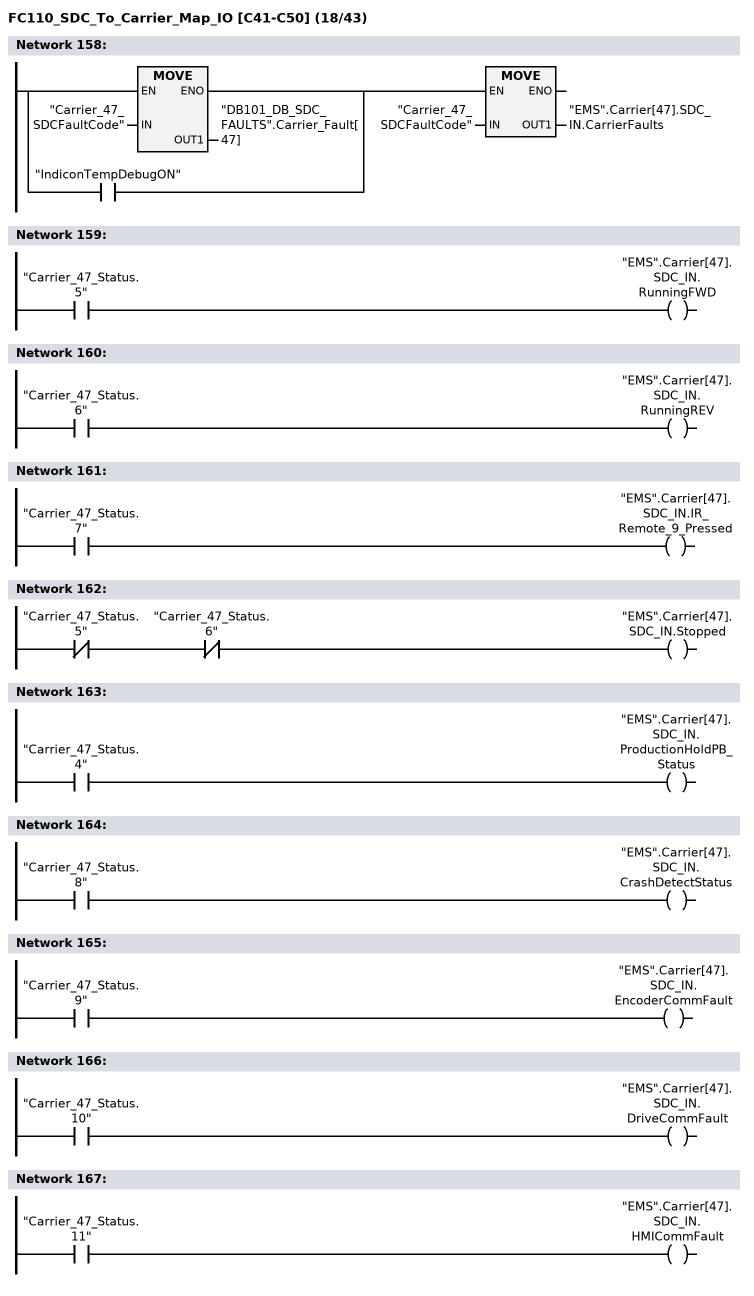
   RUNG wire#powerrail
      Move(in := "Carrier_47_SDCFaultCode", out1 => "DB101_DB_SDC_FAULTS".Carrier_Fault[47])
      wire#w1
      Move(in := "Carrier_47_SDCFaultCode", out1 => "EMS".Carrier[47].SDC_IN.CarrierFaults)
   END_RUNG
   RUNG wire#powerrail
      Contact( "IndiconTempDebugON" )
   END_RUNG wire#w1
   // the same network as SCL:
   "DB101_DB_SDC_FAULTS".Carrier_Fault[47] := "Carrier_47_SDCFaultCode";
   IF TRUE OR "IndiconTempDebugON" THEN
       "EMS".Carrier[47].SDC_IN.CarrierFaults := "Carrier_47_SDCFaultCode";
   END_IF;
END_REGION

REGION Network 159
   RUNG wire#powerrail
      Contact( "Carrier_47_Status.5" )
      Coil( "EMS".Carrier[47].SDC_IN.RunningFWD )
   END_RUNG
   // the same network as SCL:
   "EMS".Carrier[47].SDC_IN.RunningFWD := "Carrier_47_Status.5";
END_REGION

REGION Network 160
   RUNG wire#powerrail
      Contact( "Carrier_47_Status.6" )
      Coil( "EMS".Carrier[47].SDC_IN.RunningREV )
   END_RUNG
   // the same network as SCL:
   "EMS".Carrier[47].SDC_IN.RunningREV := "Carrier_47_Status.6";
END_REGION

REGION Network 161
   RUNG wire#powerrail
      Contact( "Carrier_47_Status.7" )
      Coil( "EMS".Carrier[47].SDC_IN.IR_Remote_9_Pressed )
   END_RUNG
   // the same network as SCL:
   "EMS".Carrier[47].SDC_IN.IR_Remote_9_Pressed := "Carrier_47_Status.7";
END_REGION

REGION Network 162
   RUNG wire#powerrail
      I_Contact( "Carrier_47_Status.5" )
      I_Contact( "Carrier_47_Status.6" )
      Coil( "EMS".Carrier[47].SDC_IN.Stopped )
   END_RUNG
   // the same network as SCL:
   "EMS".Carrier[47].SDC_IN.Stopped := NOT "Carrier_47_Status.5" AND NOT "Carrier_47_Status.6";
END_REGION

REGION Network 163
   RUNG wire#powerrail
      Contact( "Carrier_47_Status.4" )
      Coil( "EMS".Carrier[47].SDC_IN.ProductionHoldPB_Status )
   END_RUNG
   // the same network as SCL:
   "EMS".Carrier[47].SDC_IN.ProductionHoldPB_Status := "Carrier_47_Status.4";
END_REGION

REGION Network 164
   RUNG wire#powerrail
      Contact( "Carrier_47_Status.8" )
      Coil( "EMS".Carrier[47].SDC_IN.CrashDetectStatus )
   END_RUNG
   // the same network as SCL:
   "EMS".Carrier[47].SDC_IN.CrashDetectStatus := "Carrier_47_Status.8";
END_REGION

REGION Network 165
   RUNG wire#powerrail
      Contact( "Carrier_47_Status.9" )
      Coil( "EMS".Carrier[47].SDC_IN.EncoderCommFault )
   END_RUNG
   // the same network as SCL:
   "EMS".Carrier[47].SDC_IN.EncoderCommFault := "Carrier_47_Status.9";
END_REGION

REGION Network 166
   RUNG wire#powerrail
      Contact( "Carrier_47_Status.10" )
      Coil( "EMS".Carrier[47].SDC_IN.DriveCommFault )
   END_RUNG
   // the same network as SCL:
   "EMS".Carrier[47].SDC_IN.DriveCommFault := "Carrier_47_Status.10";
END_REGION

REGION Network 167
   RUNG wire#powerrail
      Contact( "Carrier_47_Status.11" )
      Coil( "EMS".Carrier[47].SDC_IN.HMICommFault )
   END_RUNG
   // the same network as SCL:
   "EMS".Carrier[47].SDC_IN.HMICommFault := "Carrier_47_Status.11";
END_REGION

REGION Network 168
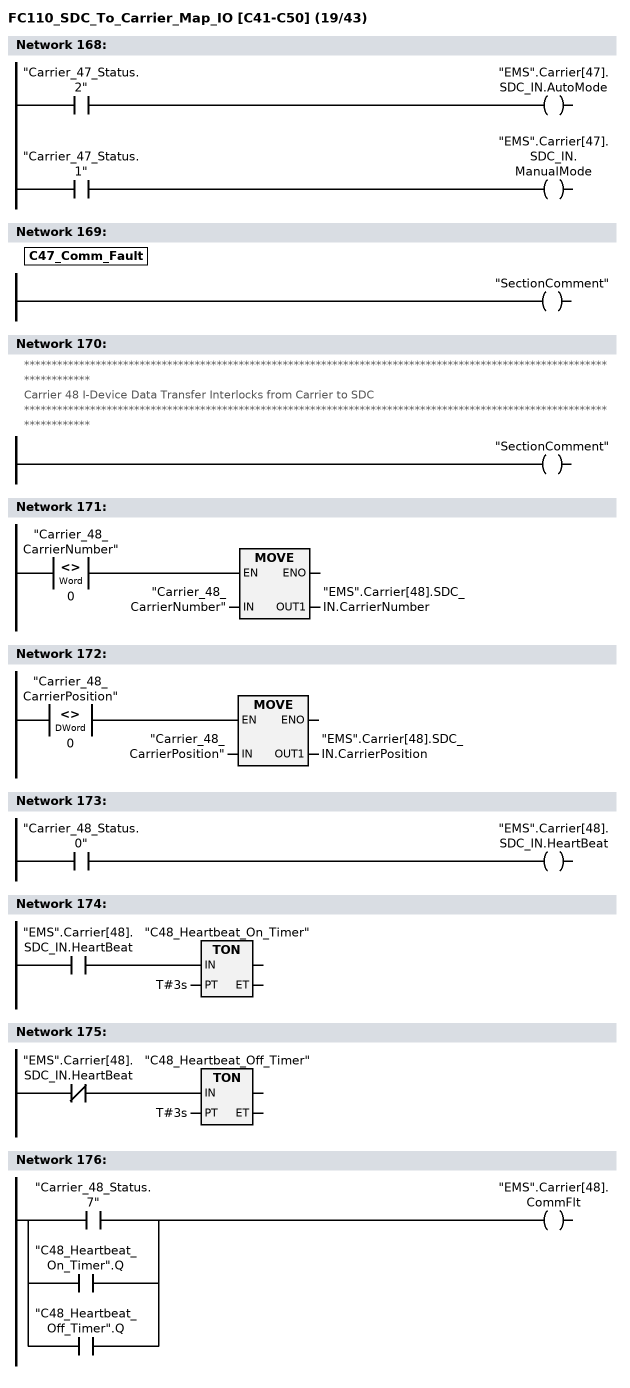
   RUNG wire#powerrail
      Contact( "Carrier_47_Status.2" )
      Coil( "EMS".Carrier[47].SDC_IN.AutoMode )
   END_RUNG
   RUNG wire#powerrail
      Contact( "Carrier_47_Status.1" )
      Coil( "EMS".Carrier[47].SDC_IN.ManualMode )
   END_RUNG
   // the same network as SCL:
   "EMS".Carrier[47].SDC_IN.AutoMode := "Carrier_47_Status.2";
   "EMS".Carrier[47].SDC_IN.ManualMode := "Carrier_47_Status.1";
END_REGION

REGION Network 169
   Label( C47_Comm_Fault )
   RUNG wire#powerrail
      Coil( "SectionComment" )
   END_RUNG
   // the same network as SCL:
   C47_Comm_Fault:
   "SectionComment" := TRUE;
END_REGION

REGION Network 170
   // **********************************************************************************************************************
   // 
   // Carrier 48 I-Device Data Transfer Interlocks from Carrier to SDC
   // 
   // **********************************************************************************************************************
   RUNG wire#powerrail
      Coil( "SectionComment" )
   END_RUNG
   // the same network as SCL:
   "SectionComment" := TRUE;
END_REGION

REGION Network 171
   RUNG wire#powerrail
      { S7_Templates := "SrcType := Word" } NE_Contact(in1 := "Carrier_48_CarrierNumber", in2 := 0)
      Move(in := "Carrier_48_CarrierNumber", out1 => "EMS".Carrier[48].SDC_IN.CarrierNumber)
   END_RUNG
   // the same network as SCL:
   IF "Carrier_48_CarrierNumber" <> 0 THEN
       "EMS".Carrier[48].SDC_IN.CarrierNumber := "Carrier_48_CarrierNumber";
   END_IF;
END_REGION

REGION Network 172
   RUNG wire#powerrail
      { S7_Templates := "SrcType := DWord" } NE_Contact(in1 := "Carrier_48_CarrierPosition", in2 := 0)
      Move(in := "Carrier_48_CarrierPosition", out1 => "EMS".Carrier[48].SDC_IN.CarrierPosition)
   END_RUNG
   // the same network as SCL:
   IF "Carrier_48_CarrierPosition" <> 0 THEN
       "EMS".Carrier[48].SDC_IN.CarrierPosition := "Carrier_48_CarrierPosition";
   END_IF;
END_REGION

REGION Network 173
   RUNG wire#powerrail
      Contact( "Carrier_48_Status.0" )
      Coil( "EMS".Carrier[48].SDC_IN.HeartBeat )
   END_RUNG
   // the same network as SCL:
   "EMS".Carrier[48].SDC_IN.HeartBeat := "Carrier_48_Status.0";
END_REGION

REGION Network 174
   "C48_Heartbeat_On_Timer".TON(IN := "EMS".Carrier[48].SDC_IN.HeartBeat, PT := T#3s);
END_REGION

REGION Network 175
   "C48_Heartbeat_Off_Timer".TON(IN := NOT "EMS".Carrier[48].SDC_IN.HeartBeat, PT := T#3s);
END_REGION

REGION Network 176
   RUNG wire#powerrail
      Contact( "Carrier_48_Status.7" )
      wire#w1
      Coil( "EMS".Carrier[48].CommFlt )
   END_RUNG
   RUNG wire#powerrail
      Contact( "C48_Heartbeat_On_Timer".Q )
   END_RUNG wire#w1
   RUNG wire#powerrail
      Contact( "C48_Heartbeat_Off_Timer".Q )
   END_RUNG wire#w1
   // the same network as SCL:
   "EMS".Carrier[48].CommFlt := "Carrier_48_Status.7" OR "C48_Heartbeat_On_Timer".Q OR "C48_Heartbeat_Off_Timer".Q;
END_REGION

REGION Network 177
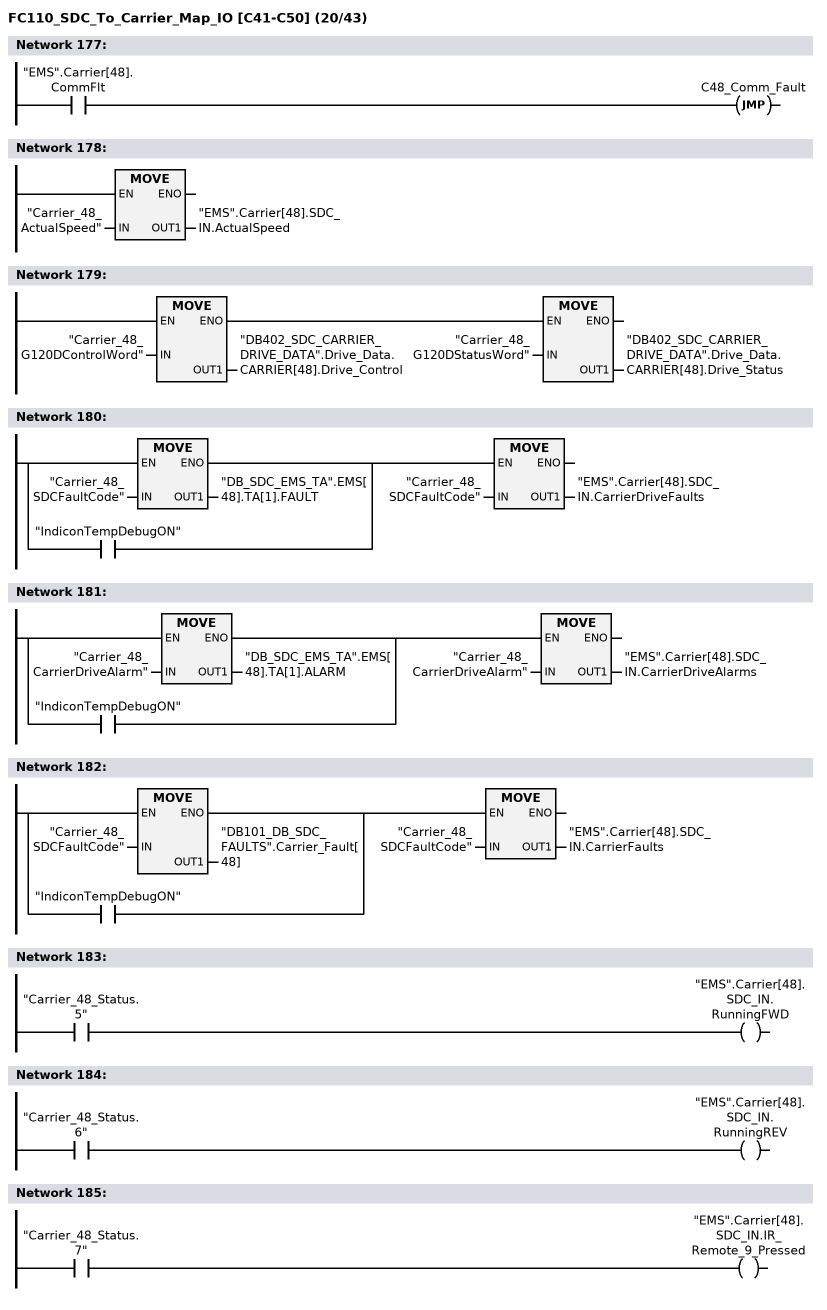
   RUNG wire#powerrail
      Contact( "EMS".Carrier[48].CommFlt )
      JumpCoil( C48_Comm_Fault )
   END_RUNG
   // the same network as SCL:
   IF "EMS".Carrier[48].CommFlt THEN GOTO C48_Comm_Fault; END_IF;
END_REGION

REGION Network 178
   RUNG wire#powerrail
      Move(in := "Carrier_48_ActualSpeed", out1 => "EMS".Carrier[48].SDC_IN.ActualSpeed)
   END_RUNG
   // the same network as SCL:
   "EMS".Carrier[48].SDC_IN.ActualSpeed := "Carrier_48_ActualSpeed";
END_REGION

REGION Network 179
   RUNG wire#powerrail
      Move(in := "Carrier_48_G120DControlWord", out1 => "DB402_SDC_CARRIER_DRIVE_DATA".Drive_Data.CARRIER[48].Drive_Control)
      Move(in := "Carrier_48_G120DStatusWord", out1 => "DB402_SDC_CARRIER_DRIVE_DATA".Drive_Data.CARRIER[48].Drive_Status)
   END_RUNG
   // the same network as SCL:
   "DB402_SDC_CARRIER_DRIVE_DATA".Drive_Data.CARRIER[48].Drive_Control := "Carrier_48_G120DControlWord";
   "DB402_SDC_CARRIER_DRIVE_DATA".Drive_Data.CARRIER[48].Drive_Status := "Carrier_48_G120DStatusWord";
END_REGION

REGION Network 180
   RUNG wire#powerrail
      Move(in := "Carrier_48_SDCFaultCode", out1 => "DB_SDC_EMS_TA".EMS[48].TA[1].FAULT)
      wire#w1
      Move(in := "Carrier_48_SDCFaultCode", out1 => "EMS".Carrier[48].SDC_IN.CarrierDriveFaults)
   END_RUNG
   RUNG wire#powerrail
      Contact( "IndiconTempDebugON" )
   END_RUNG wire#w1
   // the same network as SCL:
   "DB_SDC_EMS_TA".EMS[48].TA[1].FAULT := "Carrier_48_SDCFaultCode";
   IF TRUE OR "IndiconTempDebugON" THEN
       "EMS".Carrier[48].SDC_IN.CarrierDriveFaults := "Carrier_48_SDCFaultCode";
   END_IF;
END_REGION

REGION Network 181
   RUNG wire#powerrail
      Move(in := "Carrier_48_CarrierDriveAlarm", out1 => "DB_SDC_EMS_TA".EMS[48].TA[1].ALARM)
      wire#w1
      Move(in := "Carrier_48_CarrierDriveAlarm", out1 => "EMS".Carrier[48].SDC_IN.CarrierDriveAlarms)
   END_RUNG
   RUNG wire#powerrail
      Contact( "IndiconTempDebugON" )
   END_RUNG wire#w1
   // the same network as SCL:
   "DB_SDC_EMS_TA".EMS[48].TA[1].ALARM := "Carrier_48_CarrierDriveAlarm";
   IF TRUE OR "IndiconTempDebugON" THEN
       "EMS".Carrier[48].SDC_IN.CarrierDriveAlarms := "Carrier_48_CarrierDriveAlarm";
   END_IF;
END_REGION

REGION Network 182
   RUNG wire#powerrail
      Move(in := "Carrier_48_SDCFaultCode", out1 => "DB101_DB_SDC_FAULTS".Carrier_Fault[48])
      wire#w1
      Move(in := "Carrier_48_SDCFaultCode", out1 => "EMS".Carrier[48].SDC_IN.CarrierFaults)
   END_RUNG
   RUNG wire#powerrail
      Contact( "IndiconTempDebugON" )
   END_RUNG wire#w1
   // the same network as SCL:
   "DB101_DB_SDC_FAULTS".Carrier_Fault[48] := "Carrier_48_SDCFaultCode";
   IF TRUE OR "IndiconTempDebugON" THEN
       "EMS".Carrier[48].SDC_IN.CarrierFaults := "Carrier_48_SDCFaultCode";
   END_IF;
END_REGION

REGION Network 183
   RUNG wire#powerrail
      Contact( "Carrier_48_Status.5" )
      Coil( "EMS".Carrier[48].SDC_IN.RunningFWD )
   END_RUNG
   // the same network as SCL:
   "EMS".Carrier[48].SDC_IN.RunningFWD := "Carrier_48_Status.5";
END_REGION

REGION Network 184
   RUNG wire#powerrail
      Contact( "Carrier_48_Status.6" )
      Coil( "EMS".Carrier[48].SDC_IN.RunningREV )
   END_RUNG
   // the same network as SCL:
   "EMS".Carrier[48].SDC_IN.RunningREV := "Carrier_48_Status.6";
END_REGION

REGION Network 185
   RUNG wire#powerrail
      Contact( "Carrier_48_Status.7" )
      Coil( "EMS".Carrier[48].SDC_IN.IR_Remote_9_Pressed )
   END_RUNG
   // the same network as SCL:
   "EMS".Carrier[48].SDC_IN.IR_Remote_9_Pressed := "Carrier_48_Status.7";
END_REGION

REGION Network 186
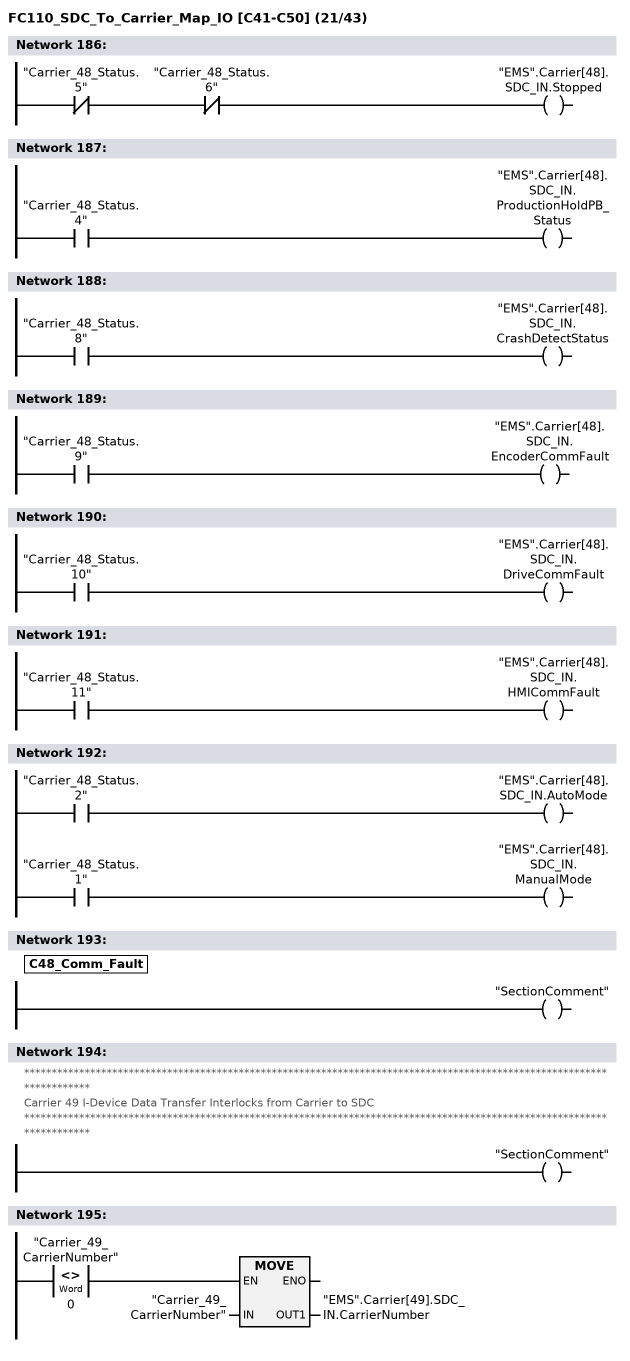
   RUNG wire#powerrail
      I_Contact( "Carrier_48_Status.5" )
      I_Contact( "Carrier_48_Status.6" )
      Coil( "EMS".Carrier[48].SDC_IN.Stopped )
   END_RUNG
   // the same network as SCL:
   "EMS".Carrier[48].SDC_IN.Stopped := NOT "Carrier_48_Status.5" AND NOT "Carrier_48_Status.6";
END_REGION

REGION Network 187
   RUNG wire#powerrail
      Contact( "Carrier_48_Status.4" )
      Coil( "EMS".Carrier[48].SDC_IN.ProductionHoldPB_Status )
   END_RUNG
   // the same network as SCL:
   "EMS".Carrier[48].SDC_IN.ProductionHoldPB_Status := "Carrier_48_Status.4";
END_REGION

REGION Network 188
   RUNG wire#powerrail
      Contact( "Carrier_48_Status.8" )
      Coil( "EMS".Carrier[48].SDC_IN.CrashDetectStatus )
   END_RUNG
   // the same network as SCL:
   "EMS".Carrier[48].SDC_IN.CrashDetectStatus := "Carrier_48_Status.8";
END_REGION

REGION Network 189
   RUNG wire#powerrail
      Contact( "Carrier_48_Status.9" )
      Coil( "EMS".Carrier[48].SDC_IN.EncoderCommFault )
   END_RUNG
   // the same network as SCL:
   "EMS".Carrier[48].SDC_IN.EncoderCommFault := "Carrier_48_Status.9";
END_REGION

REGION Network 190
   RUNG wire#powerrail
      Contact( "Carrier_48_Status.10" )
      Coil( "EMS".Carrier[48].SDC_IN.DriveCommFault )
   END_RUNG
   // the same network as SCL:
   "EMS".Carrier[48].SDC_IN.DriveCommFault := "Carrier_48_Status.10";
END_REGION

REGION Network 191
   RUNG wire#powerrail
      Contact( "Carrier_48_Status.11" )
      Coil( "EMS".Carrier[48].SDC_IN.HMICommFault )
   END_RUNG
   // the same network as SCL:
   "EMS".Carrier[48].SDC_IN.HMICommFault := "Carrier_48_Status.11";
END_REGION

REGION Network 192
   RUNG wire#powerrail
      Contact( "Carrier_48_Status.2" )
      Coil( "EMS".Carrier[48].SDC_IN.AutoMode )
   END_RUNG
   RUNG wire#powerrail
      Contact( "Carrier_48_Status.1" )
      Coil( "EMS".Carrier[48].SDC_IN.ManualMode )
   END_RUNG
   // the same network as SCL:
   "EMS".Carrier[48].SDC_IN.AutoMode := "Carrier_48_Status.2";
   "EMS".Carrier[48].SDC_IN.ManualMode := "Carrier_48_Status.1";
END_REGION

REGION Network 193
   Label( C48_Comm_Fault )
   RUNG wire#powerrail
      Coil( "SectionComment" )
   END_RUNG
   // the same network as SCL:
   C48_Comm_Fault:
   "SectionComment" := TRUE;
END_REGION

REGION Network 194
   // **********************************************************************************************************************
   // 
   // Carrier 49 I-Device Data Transfer Interlocks from Carrier to SDC
   // 
   // **********************************************************************************************************************
   RUNG wire#powerrail
      Coil( "SectionComment" )
   END_RUNG
   // the same network as SCL:
   "SectionComment" := TRUE;
END_REGION

REGION Network 195
   RUNG wire#powerrail
      { S7_Templates := "SrcType := Word" } NE_Contact(in1 := "Carrier_49_CarrierNumber", in2 := 0)
      Move(in := "Carrier_49_CarrierNumber", out1 => "EMS".Carrier[49].SDC_IN.CarrierNumber)
   END_RUNG
   // the same network as SCL:
   IF "Carrier_49_CarrierNumber" <> 0 THEN
       "EMS".Carrier[49].SDC_IN.CarrierNumber := "Carrier_49_CarrierNumber";
   END_IF;
END_REGION

REGION Network 196
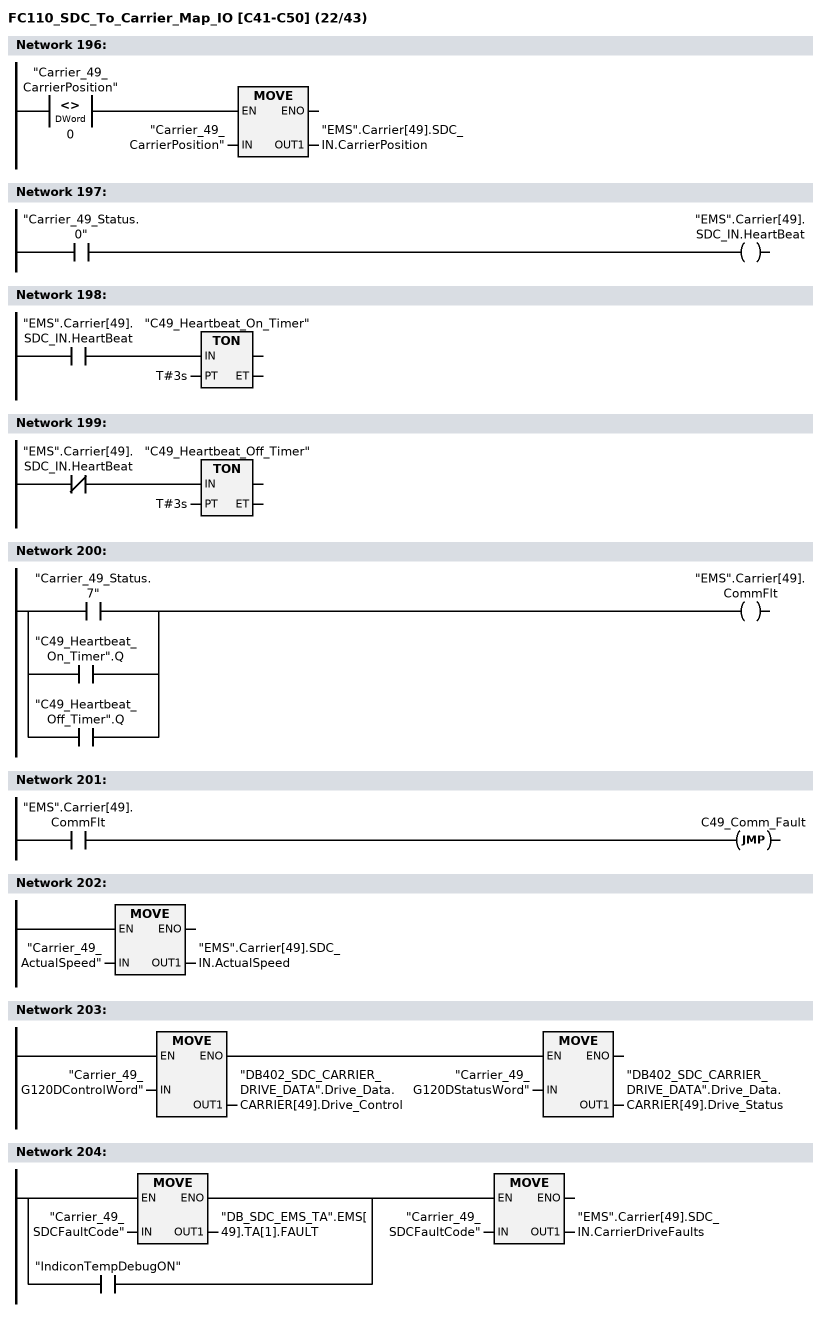
   RUNG wire#powerrail
      { S7_Templates := "SrcType := DWord" } NE_Contact(in1 := "Carrier_49_CarrierPosition", in2 := 0)
      Move(in := "Carrier_49_CarrierPosition", out1 => "EMS".Carrier[49].SDC_IN.CarrierPosition)
   END_RUNG
   // the same network as SCL:
   IF "Carrier_49_CarrierPosition" <> 0 THEN
       "EMS".Carrier[49].SDC_IN.CarrierPosition := "Carrier_49_CarrierPosition";
   END_IF;
END_REGION

REGION Network 197
   RUNG wire#powerrail
      Contact( "Carrier_49_Status.0" )
      Coil( "EMS".Carrier[49].SDC_IN.HeartBeat )
   END_RUNG
   // the same network as SCL:
   "EMS".Carrier[49].SDC_IN.HeartBeat := "Carrier_49_Status.0";
END_REGION

REGION Network 198
   "C49_Heartbeat_On_Timer".TON(IN := "EMS".Carrier[49].SDC_IN.HeartBeat, PT := T#3s);
END_REGION

REGION Network 199
   "C49_Heartbeat_Off_Timer".TON(IN := NOT "EMS".Carrier[49].SDC_IN.HeartBeat, PT := T#3s);
END_REGION

REGION Network 200
   RUNG wire#powerrail
      Contact( "Carrier_49_Status.7" )
      wire#w1
      Coil( "EMS".Carrier[49].CommFlt )
   END_RUNG
   RUNG wire#powerrail
      Contact( "C49_Heartbeat_On_Timer".Q )
   END_RUNG wire#w1
   RUNG wire#powerrail
      Contact( "C49_Heartbeat_Off_Timer".Q )
   END_RUNG wire#w1
   // the same network as SCL:
   "EMS".Carrier[49].CommFlt := "Carrier_49_Status.7" OR "C49_Heartbeat_On_Timer".Q OR "C49_Heartbeat_Off_Timer".Q;
END_REGION

REGION Network 201
   RUNG wire#powerrail
      Contact( "EMS".Carrier[49].CommFlt )
      JumpCoil( C49_Comm_Fault )
   END_RUNG
   // the same network as SCL:
   IF "EMS".Carrier[49].CommFlt THEN GOTO C49_Comm_Fault; END_IF;
END_REGION

REGION Network 202
   RUNG wire#powerrail
      Move(in := "Carrier_49_ActualSpeed", out1 => "EMS".Carrier[49].SDC_IN.ActualSpeed)
   END_RUNG
   // the same network as SCL:
   "EMS".Carrier[49].SDC_IN.ActualSpeed := "Carrier_49_ActualSpeed";
END_REGION

REGION Network 203
   RUNG wire#powerrail
      Move(in := "Carrier_49_G120DControlWord", out1 => "DB402_SDC_CARRIER_DRIVE_DATA".Drive_Data.CARRIER[49].Drive_Control)
      Move(in := "Carrier_49_G120DStatusWord", out1 => "DB402_SDC_CARRIER_DRIVE_DATA".Drive_Data.CARRIER[49].Drive_Status)
   END_RUNG
   // the same network as SCL:
   "DB402_SDC_CARRIER_DRIVE_DATA".Drive_Data.CARRIER[49].Drive_Control := "Carrier_49_G120DControlWord";
   "DB402_SDC_CARRIER_DRIVE_DATA".Drive_Data.CARRIER[49].Drive_Status := "Carrier_49_G120DStatusWord";
END_REGION

REGION Network 204
   RUNG wire#powerrail
      Move(in := "Carrier_49_SDCFaultCode", out1 => "DB_SDC_EMS_TA".EMS[49].TA[1].FAULT)
      wire#w1
      Move(in := "Carrier_49_SDCFaultCode", out1 => "EMS".Carrier[49].SDC_IN.CarrierDriveFaults)
   END_RUNG
   RUNG wire#powerrail
      Contact( "IndiconTempDebugON" )
   END_RUNG wire#w1
   // the same network as SCL:
   "DB_SDC_EMS_TA".EMS[49].TA[1].FAULT := "Carrier_49_SDCFaultCode";
   IF TRUE OR "IndiconTempDebugON" THEN
       "EMS".Carrier[49].SDC_IN.CarrierDriveFaults := "Carrier_49_SDCFaultCode";
   END_IF;
END_REGION

REGION Network 205
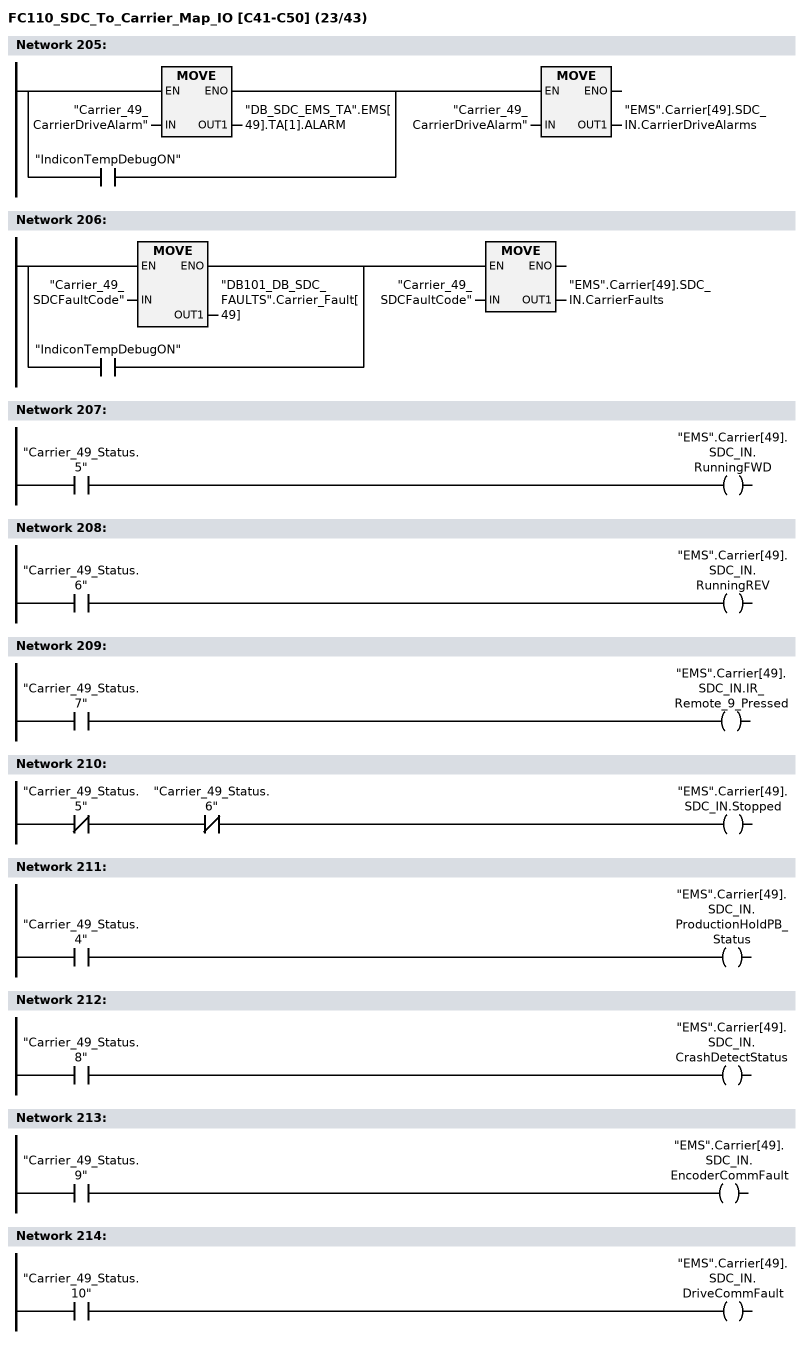
   RUNG wire#powerrail
      Move(in := "Carrier_49_CarrierDriveAlarm", out1 => "DB_SDC_EMS_TA".EMS[49].TA[1].ALARM)
      wire#w1
      Move(in := "Carrier_49_CarrierDriveAlarm", out1 => "EMS".Carrier[49].SDC_IN.CarrierDriveAlarms)
   END_RUNG
   RUNG wire#powerrail
      Contact( "IndiconTempDebugON" )
   END_RUNG wire#w1
   // the same network as SCL:
   "DB_SDC_EMS_TA".EMS[49].TA[1].ALARM := "Carrier_49_CarrierDriveAlarm";
   IF TRUE OR "IndiconTempDebugON" THEN
       "EMS".Carrier[49].SDC_IN.CarrierDriveAlarms := "Carrier_49_CarrierDriveAlarm";
   END_IF;
END_REGION

REGION Network 206
   RUNG wire#powerrail
      Move(in := "Carrier_49_SDCFaultCode", out1 => "DB101_DB_SDC_FAULTS".Carrier_Fault[49])
      wire#w1
      Move(in := "Carrier_49_SDCFaultCode", out1 => "EMS".Carrier[49].SDC_IN.CarrierFaults)
   END_RUNG
   RUNG wire#powerrail
      Contact( "IndiconTempDebugON" )
   END_RUNG wire#w1
   // the same network as SCL:
   "DB101_DB_SDC_FAULTS".Carrier_Fault[49] := "Carrier_49_SDCFaultCode";
   IF TRUE OR "IndiconTempDebugON" THEN
       "EMS".Carrier[49].SDC_IN.CarrierFaults := "Carrier_49_SDCFaultCode";
   END_IF;
END_REGION

REGION Network 207
   RUNG wire#powerrail
      Contact( "Carrier_49_Status.5" )
      Coil( "EMS".Carrier[49].SDC_IN.RunningFWD )
   END_RUNG
   // the same network as SCL:
   "EMS".Carrier[49].SDC_IN.RunningFWD := "Carrier_49_Status.5";
END_REGION

REGION Network 208
   RUNG wire#powerrail
      Contact( "Carrier_49_Status.6" )
      Coil( "EMS".Carrier[49].SDC_IN.RunningREV )
   END_RUNG
   // the same network as SCL:
   "EMS".Carrier[49].SDC_IN.RunningREV := "Carrier_49_Status.6";
END_REGION

REGION Network 209
   RUNG wire#powerrail
      Contact( "Carrier_49_Status.7" )
      Coil( "EMS".Carrier[49].SDC_IN.IR_Remote_9_Pressed )
   END_RUNG
   // the same network as SCL:
   "EMS".Carrier[49].SDC_IN.IR_Remote_9_Pressed := "Carrier_49_Status.7";
END_REGION

REGION Network 210
   RUNG wire#powerrail
      I_Contact( "Carrier_49_Status.5" )
      I_Contact( "Carrier_49_Status.6" )
      Coil( "EMS".Carrier[49].SDC_IN.Stopped )
   END_RUNG
   // the same network as SCL:
   "EMS".Carrier[49].SDC_IN.Stopped := NOT "Carrier_49_Status.5" AND NOT "Carrier_49_Status.6";
END_REGION

REGION Network 211
   RUNG wire#powerrail
      Contact( "Carrier_49_Status.4" )
      Coil( "EMS".Carrier[49].SDC_IN.ProductionHoldPB_Status )
   END_RUNG
   // the same network as SCL:
   "EMS".Carrier[49].SDC_IN.ProductionHoldPB_Status := "Carrier_49_Status.4";
END_REGION

REGION Network 212
   RUNG wire#powerrail
      Contact( "Carrier_49_Status.8" )
      Coil( "EMS".Carrier[49].SDC_IN.CrashDetectStatus )
   END_RUNG
   // the same network as SCL:
   "EMS".Carrier[49].SDC_IN.CrashDetectStatus := "Carrier_49_Status.8";
END_REGION

REGION Network 213
   RUNG wire#powerrail
      Contact( "Carrier_49_Status.9" )
      Coil( "EMS".Carrier[49].SDC_IN.EncoderCommFault )
   END_RUNG
   // the same network as SCL:
   "EMS".Carrier[49].SDC_IN.EncoderCommFault := "Carrier_49_Status.9";
END_REGION

REGION Network 214
   RUNG wire#powerrail
      Contact( "Carrier_49_Status.10" )
      Coil( "EMS".Carrier[49].SDC_IN.DriveCommFault )
   END_RUNG
   // the same network as SCL:
   "EMS".Carrier[49].SDC_IN.DriveCommFault := "Carrier_49_Status.10";
END_REGION

REGION Network 215
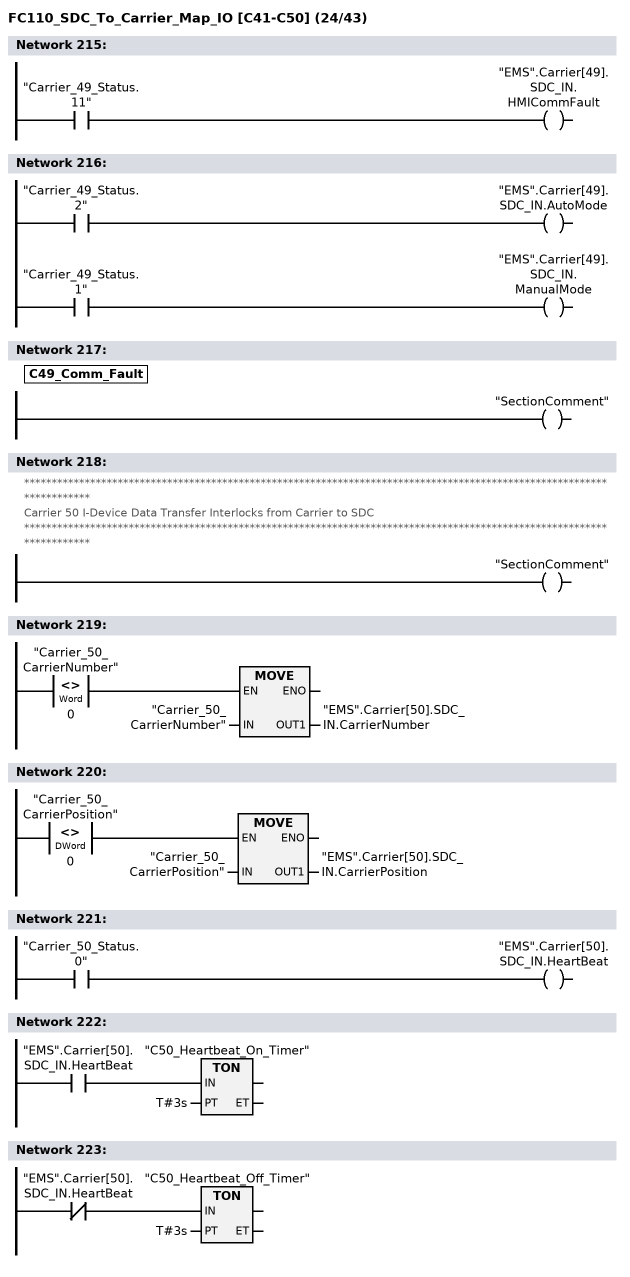
   RUNG wire#powerrail
      Contact( "Carrier_49_Status.11" )
      Coil( "EMS".Carrier[49].SDC_IN.HMICommFault )
   END_RUNG
   // the same network as SCL:
   "EMS".Carrier[49].SDC_IN.HMICommFault := "Carrier_49_Status.11";
END_REGION

REGION Network 216
   RUNG wire#powerrail
      Contact( "Carrier_49_Status.2" )
      Coil( "EMS".Carrier[49].SDC_IN.AutoMode )
   END_RUNG
   RUNG wire#powerrail
      Contact( "Carrier_49_Status.1" )
      Coil( "EMS".Carrier[49].SDC_IN.ManualMode )
   END_RUNG
   // the same network as SCL:
   "EMS".Carrier[49].SDC_IN.AutoMode := "Carrier_49_Status.2";
   "EMS".Carrier[49].SDC_IN.ManualMode := "Carrier_49_Status.1";
END_REGION

REGION Network 217
   Label( C49_Comm_Fault )
   RUNG wire#powerrail
      Coil( "SectionComment" )
   END_RUNG
   // the same network as SCL:
   C49_Comm_Fault:
   "SectionComment" := TRUE;
END_REGION

REGION Network 218
   // **********************************************************************************************************************
   // 
   // Carrier 50 I-Device Data Transfer Interlocks from Carrier to SDC
   // 
   // **********************************************************************************************************************
   RUNG wire#powerrail
      Coil( "SectionComment" )
   END_RUNG
   // the same network as SCL:
   "SectionComment" := TRUE;
END_REGION

REGION Network 219
   RUNG wire#powerrail
      { S7_Templates := "SrcType := Word" } NE_Contact(in1 := "Carrier_50_CarrierNumber", in2 := 0)
      Move(in := "Carrier_50_CarrierNumber", out1 => "EMS".Carrier[50].SDC_IN.CarrierNumber)
   END_RUNG
   // the same network as SCL:
   IF "Carrier_50_CarrierNumber" <> 0 THEN
       "EMS".Carrier[50].SDC_IN.CarrierNumber := "Carrier_50_CarrierNumber";
   END_IF;
END_REGION

REGION Network 220
   RUNG wire#powerrail
      { S7_Templates := "SrcType := DWord" } NE_Contact(in1 := "Carrier_50_CarrierPosition", in2 := 0)
      Move(in := "Carrier_50_CarrierPosition", out1 => "EMS".Carrier[50].SDC_IN.CarrierPosition)
   END_RUNG
   // the same network as SCL:
   IF "Carrier_50_CarrierPosition" <> 0 THEN
       "EMS".Carrier[50].SDC_IN.CarrierPosition := "Carrier_50_CarrierPosition";
   END_IF;
END_REGION

REGION Network 221
   RUNG wire#powerrail
      Contact( "Carrier_50_Status.0" )
      Coil( "EMS".Carrier[50].SDC_IN.HeartBeat )
   END_RUNG
   // the same network as SCL:
   "EMS".Carrier[50].SDC_IN.HeartBeat := "Carrier_50_Status.0";
END_REGION

REGION Network 222
   "C50_Heartbeat_On_Timer".TON(IN := "EMS".Carrier[50].SDC_IN.HeartBeat, PT := T#3s);
END_REGION

REGION Network 223
   "C50_Heartbeat_Off_Timer".TON(IN := NOT "EMS".Carrier[50].SDC_IN.HeartBeat, PT := T#3s);
END_REGION

REGION Network 224